(* Logix 5000 project; controller PLC_MCC1300_75F1 vendor 1 type 14 code 166 rev 32.11; software revision 32.04; part 43 of 83 *)
(* tags used below, declared in another part *)
   AUX_xDebugNewPlate : BOOL;
   CM_INPUT_Z200_Sync : CM_INPUT_Z200;
   CONST_tAux : AUX_COSTANTS;
   CONST_tPlant : UDT_PLANT_CONSTANTS;
   GP_AccTimeForGap : GP_AccTimeForGap;
   GP_TrackingAddCap : GP_TrackingAddCap;
   GP_TrackingSearchPlate : GP_TrackingSearchPlate;
   M302SpeedUp : MAC_SpeedUp;
   M302SpeedUp_ALM : MAC_SpeedUp_ALM;
   M302SpeedUp_HMR : MAC_SpeedUp_HMR;
   M302SpeedUp_tmON_ProtSnap : TIMER;
   M302SpeedUp_xFirstScanProtSnap : BOOL;
   TMP_d : DINT;
   TMP_dDebug : DINT;
   TMP_dIndex : DINT;
   TMP_dLehrSpeed : DINT;
   TMP_x : BOOL;
   xAlwaysOFF : BOOL;
   xDebugOFF : BOOL;
   Z200_SnapDataEth : UDT_ConvoyCap_ZC[2];
   Z300_BufferPlate : UDT_LINE_BUFFER_PLATE;
   Z300_Conveyor : UDT_StandConv[29];
   Z300_dEndTrackingPosition : DINT;
   Z300_LineTracking : UDT_LINE_TRACKING;
   Z301 : MAC_Zone_ML;
   Z301_HMR : MAC_Zone_ML_HMR;
(* MainProgram, continued *)

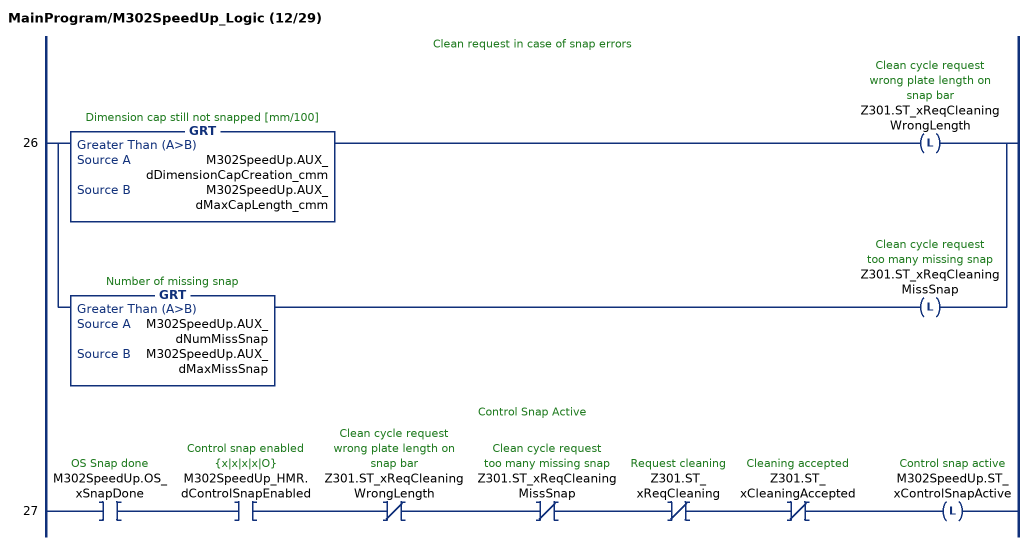
   [picture p613: MainProgram/M302SpeedUp_Logic rungs 26-27]
   // Clean request in case of snap errors
   26: [GRT(M302SpeedUp.AUX_dDimensionCapCreation_cmm,M302SpeedUp.AUX_dMaxCapLength_cmm) OTL(Z301.ST_xReqCleaningWrongLength) ,GRT(M302SpeedUp.AUX_dNumMissSnap,M302SpeedUp.AUX_dMaxMissSnap) OTL(Z301.ST_xReqCleaningMissSnap) ];
   // Control Snap Active
   27: XIC(M302SpeedUp.OS_xSnapDone)XIC(M302SpeedUp_HMR.dControlSnapEnabled)XIO(Z301.ST_xReqCleaningWrongLength)XIO(Z301.ST_xReqCleaningMissSnap)XIO(Z301.ST_xReqCleaning)XIO(Z301.ST_xCleaningAccepted)OTL(M302SpeedUp.ST_xControlSnapActive);
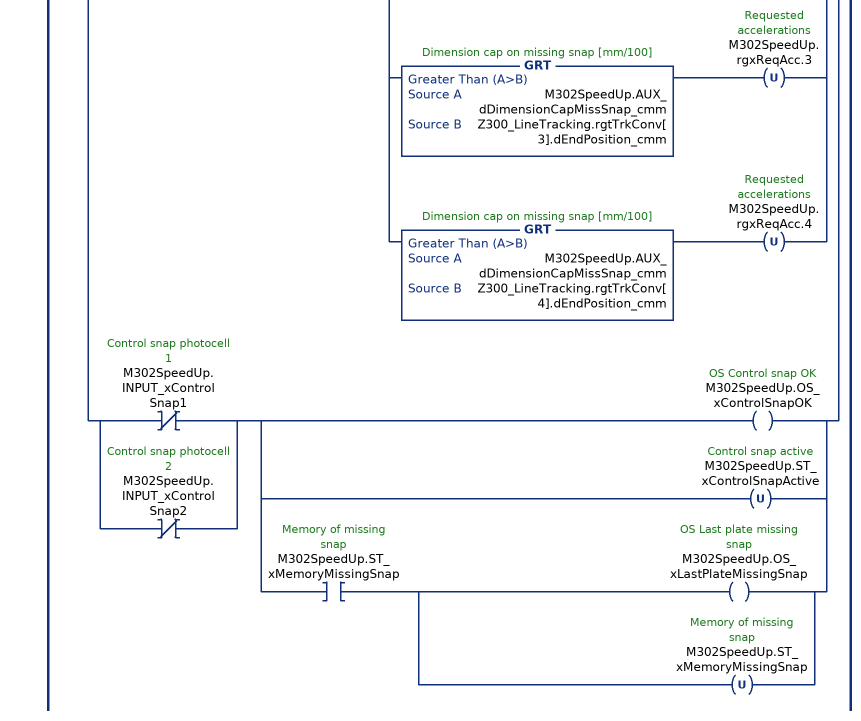
   // Missing Snap
   28: XIC(M302SpeedUp.ST_xControlSnapActive)MOV(30000,M302SpeedUp.AUX_dControlSnapLimit_cmm)[GRT(M302SpeedUp.AUX_dDimensionCapCreation_cmm,M302SpeedUp.AUX_dControlSnapLimit_cmm) [OTE(M302SpeedUp.OS_xMissingSnap) ,OTU(M302SpeedUp.ST_xControlSnapActive) ,OTU(M302SpeedUp.xReqAccAll) ,OTL(M302SpeedUp.ST_xMemoryMissingSnap) ,GRT(M302SpeedUp.AUX_dDimensionCapMissSnap_cmm,Z300_LineTracking.rgtTrkConv[0].dEndPosition_cmm) OTU(M302SpeedUp.rgxReqAcc.0) ,GRT(M302SpeedUp.AUX_dDimensionCapMissSnap_cmm,Z300_LineTracking.rgtTrkConv[1].dEndPosition_cmm) OTU(M302SpeedUp.rgxReqAcc.1) ,GRT(M302SpeedUp.AUX_dDimensionCapMissSnap_cmm,Z300_LineTracking.rgtTrkConv[2].dEndPosition_cmm) OTU(M302SpeedUp.rgxReqAcc.2) ,GRT(M302SpeedUp.AUX_dDimensionCapMissSnap_cmm,Z300_LineTracking.rgtTrkConv[3].dEndPosition_cmm) OTU(M302SpeedUp.rgxReqAcc.3) ,GRT(M302SpeedUp.AUX_dDimensionCapMissSnap_cmm,Z300_LineTracking.rgtTrkConv[4].dEndPosition_cmm) OTU(M302SpeedUp.rgxReqAcc.4) ] ,[XIO(M302SpeedUp.INPUT_xControlSnap1) ,XIO(M302SpeedUp.INPUT_xControlSnap2) ] [OTE(M302SpeedUp.OS_xControlSnapOK) ,OTU(M302SpeedUp.ST_xControlSnapActive) ,XIC(M302SpeedUp.ST_xMemoryMissingSnap) [OTE(M302SpeedUp.OS_xLastPlateMissingSnap) ,OTU(M302SpeedUp.ST_xMemoryMissingSnap) ] ] ];
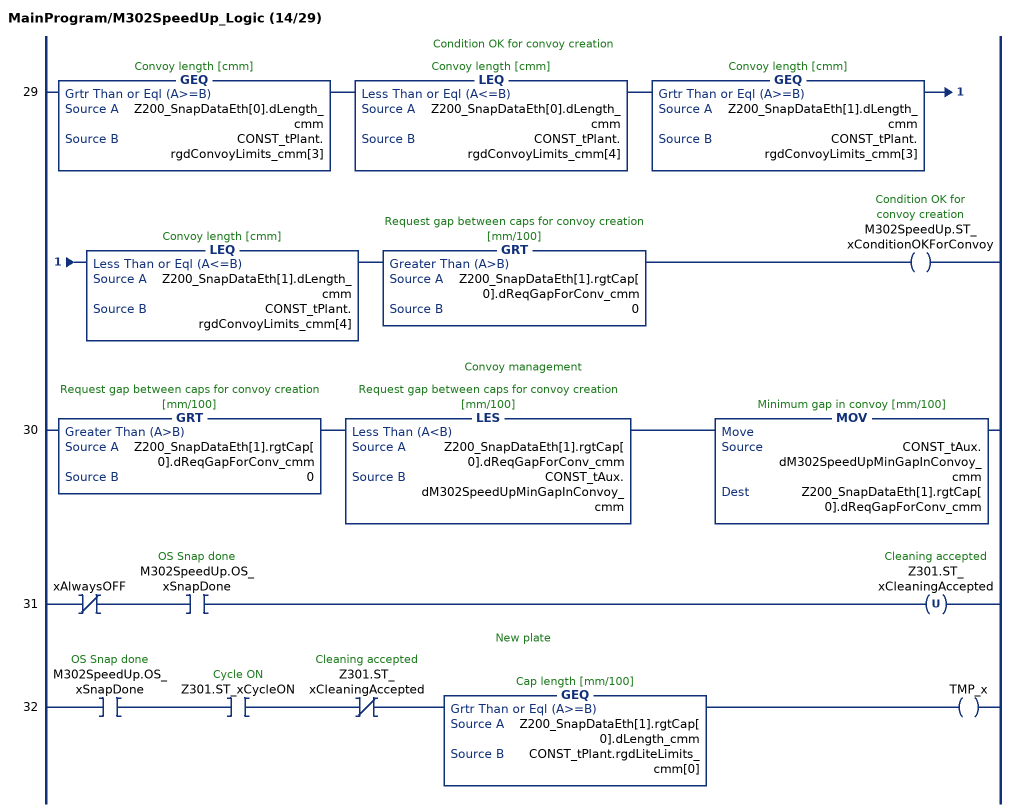
   // Condition OK for convoy creation
   29: GEQ(Z200_SnapDataEth[0].dLength_cmm,CONST_tPlant.rgdConvoyLimits_cmm[3])LEQ(Z200_SnapDataEth[0].dLength_cmm,CONST_tPlant.rgdConvoyLimits_cmm[4])GEQ(Z200_SnapDataEth[1].dLength_cmm,CONST_tPlant.rgdConvoyLimits_cmm[3])LEQ(Z200_SnapDataEth[1].dLength_cmm,CONST_tPlant.rgdConvoyLimits_cmm[4])GRT(Z200_SnapDataEth[1].rgtCap[0].dReqGapForConv_cmm,0)OTE(M302SpeedUp.ST_xConditionOKForConvoy);
   // Convoy management
   30: GRT(Z200_SnapDataEth[1].rgtCap[0].dReqGapForConv_cmm,0)LES(Z200_SnapDataEth[1].rgtCap[0].dReqGapForConv_cmm,CONST_tAux.dM302SpeedUpMinGapInConvoy_cmm)MOV(CONST_tAux.dM302SpeedUpMinGapInConvoy_cmm,Z200_SnapDataEth[1].rgtCap[0].dReqGapForConv_cmm);
   31: XIO(xAlwaysOFF)XIC(M302SpeedUp.OS_xSnapDone)OTU(Z301.ST_xCleaningAccepted);
   // New plate
   32: XIC(M302SpeedUp.OS_xSnapDone)XIC(Z301.ST_xCycleON)XIO(Z301.ST_xCleaningAccepted)GEQ(Z200_SnapDataEth[1].rgtCap[0].dLength_cmm,CONST_tPlant.rgdLiteLimits_cmm[0])OTE(TMP_x);
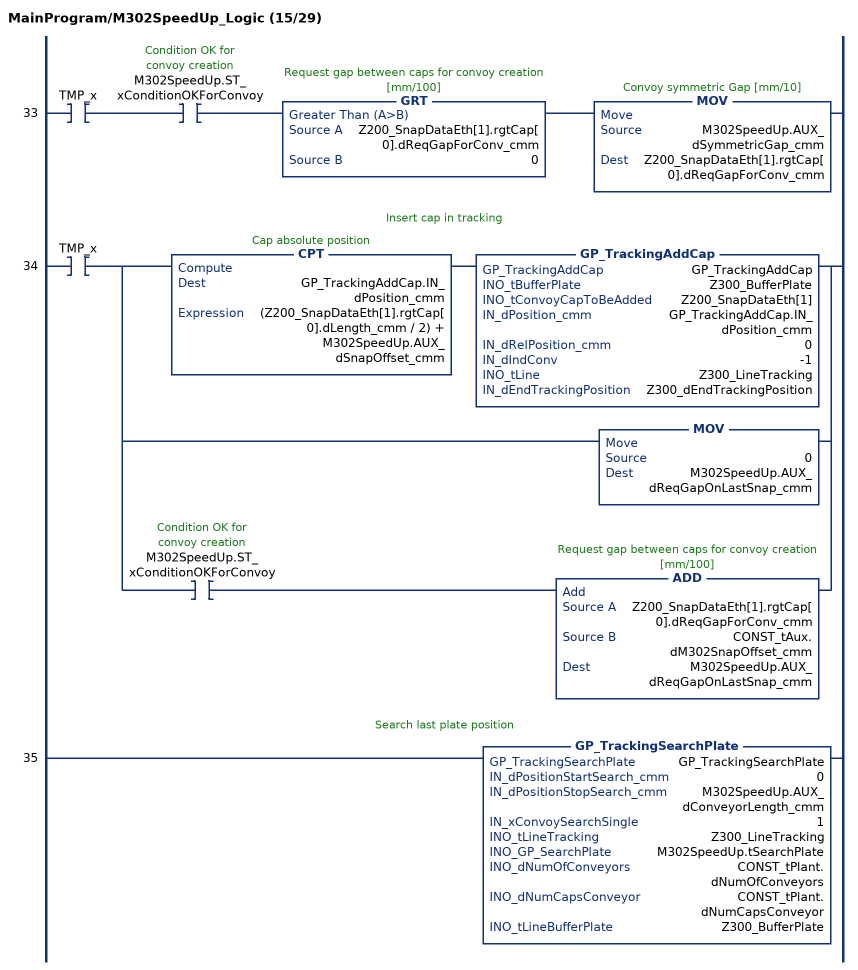
   33: XIC(TMP_x)XIC(M302SpeedUp.ST_xConditionOKForConvoy)GRT(Z200_SnapDataEth[1].rgtCap[0].dReqGapForConv_cmm,0)MOV(M302SpeedUp.AUX_dSymmetricGap_cmm,Z200_SnapDataEth[1].rgtCap[0].dReqGapForConv_cmm);
   // Insert cap in tracking
   34: XIC(TMP_x)[CPT(GP_TrackingAddCap.IN_dPosition_cmm,(Z200_SnapDataEth[1].rgtCap[0].dLength_cmm / 2) + M302SpeedUp.AUX_dSnapOffset_cmm) GP_TrackingAddCap(GP_TrackingAddCap,Z300_BufferPlate,Z200_SnapDataEth[1],GP_TrackingAddCap.IN_dPosition_cmm,0,-1,Z300_LineTracking,Z300_dEndTrackingPosition) ,MOV(0,M302SpeedUp.AUX_dReqGapOnLastSnap_cmm) ,XIC(M302SpeedUp.ST_xConditionOKForConvoy) ADD(Z200_SnapDataEth[1].rgtCap[0].dReqGapForConv_cmm,CONST_tAux.dM302SnapOffset_cmm,M302SpeedUp.AUX_dReqGapOnLastSnap_cmm) ];
   // Search last plate position
   35: GP_TrackingSearchPlate(GP_TrackingSearchPlate,0,M302SpeedUp.AUX_dConveyorLength_cmm,1,Z300_LineTracking,M302SpeedUp.tSearchPlate,CONST_tPlant.dNumOfConveyors,CONST_tPlant.dNumCapsConveyor,Z300_BufferPlate);
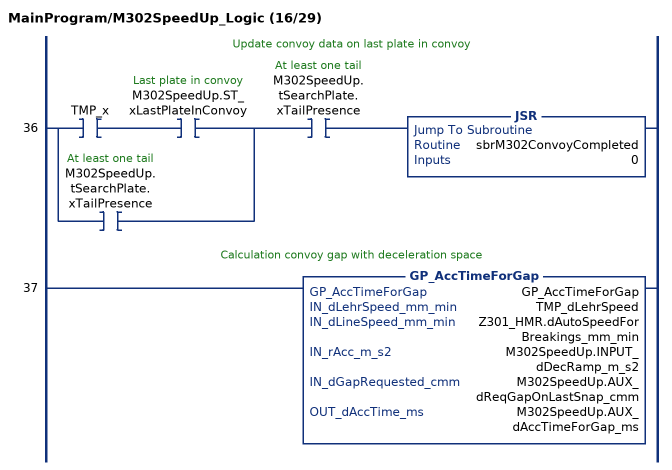
   // Update convoy data on last plate in convoy
   36: [XIC(TMP_x) XIC(M302SpeedUp.ST_xLastPlateInConvoy) ,XIC(M302SpeedUp.tSearchPlate.xTailPresence) ]XIC(M302SpeedUp.tSearchPlate.xTailPresence)JSR(sbrM302ConvoyCompleted,0);
   // Calculation convoy gap with deceleration space
   37: GP_AccTimeForGap(GP_AccTimeForGap,TMP_dLehrSpeed,Z301_HMR.dAutoSpeedForBreakings_mm_min,M302SpeedUp.INPUT_dDecRamp_m_s2,M302SpeedUp.AUX_dReqGapOnLastSnap_cmm,M302SpeedUp.AUX_dAccTimeForGap_ms);
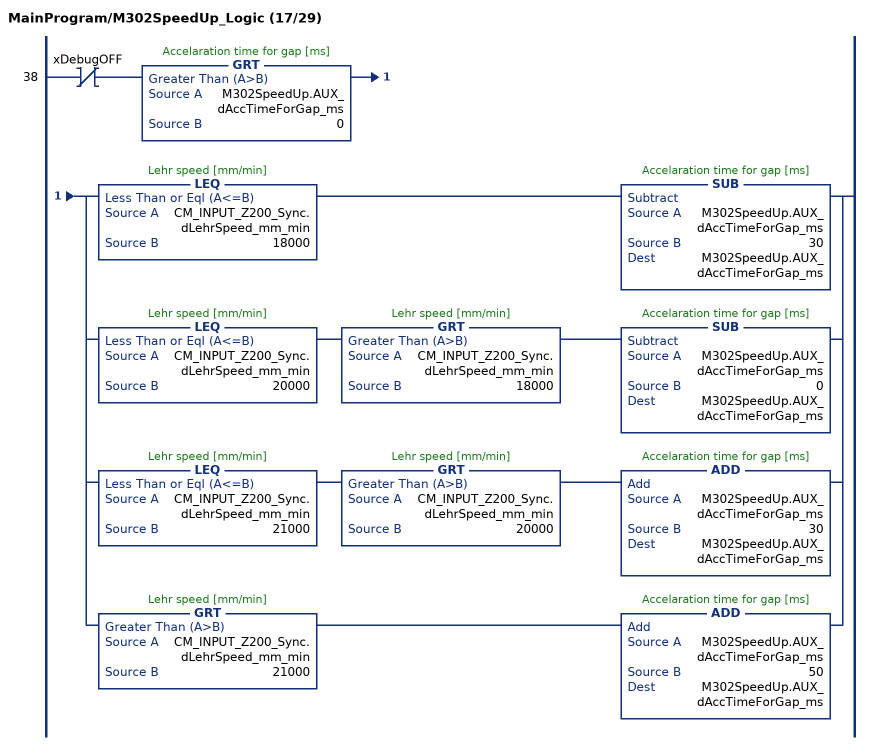
   38: XIO(xDebugOFF)GRT(M302SpeedUp.AUX_dAccTimeForGap_ms,0)[LEQ(CM_INPUT_Z200_Sync.dLehrSpeed_mm_min,18000) SUB(M302SpeedUp.AUX_dAccTimeForGap_ms,30,M302SpeedUp.AUX_dAccTimeForGap_ms) ,LEQ(CM_INPUT_Z200_Sync.dLehrSpeed_mm_min,20000) GRT(CM_INPUT_Z200_Sync.dLehrSpeed_mm_min,18000) SUB(M302SpeedUp.AUX_dAccTimeForGap_ms,0,M302SpeedUp.AUX_dAccTimeForGap_ms) ,LEQ(CM_INPUT_Z200_Sync.dLehrSpeed_mm_min,21000) GRT(CM_INPUT_Z200_Sync.dLehrSpeed_mm_min,20000) ADD(M302SpeedUp.AUX_dAccTimeForGap_ms,30,M302SpeedUp.AUX_dAccTimeForGap_ms) ,GRT(CM_INPUT_Z200_Sync.dLehrSpeed_mm_min,21000) ADD(M302SpeedUp.AUX_dAccTimeForGap_ms,50,M302SpeedUp.AUX_dAccTimeForGap_ms) ];
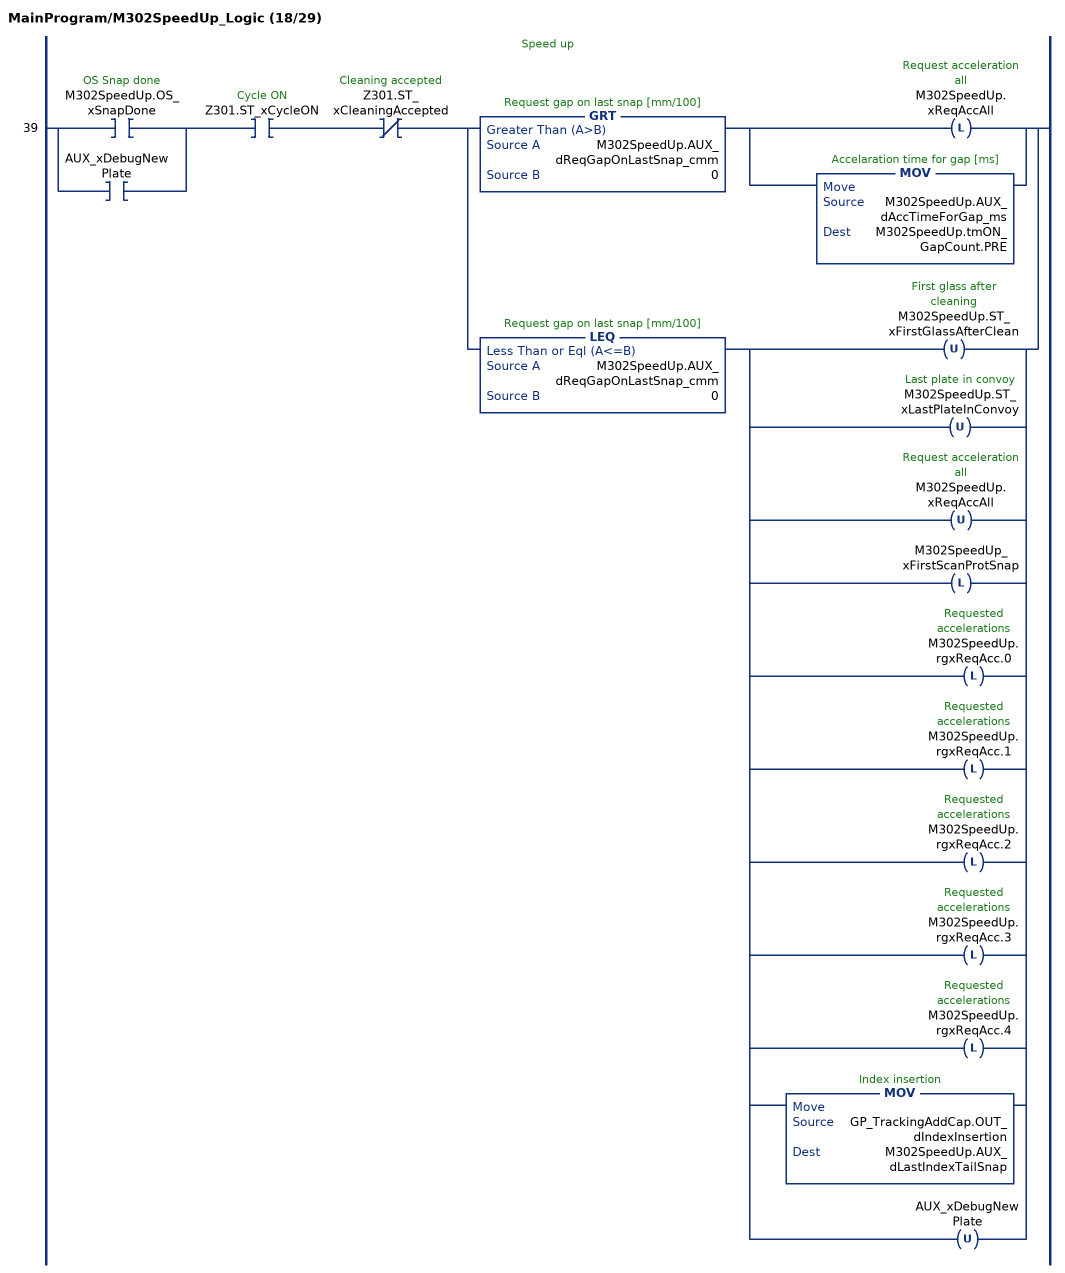
   // Speed up
   39: [XIC(M302SpeedUp.OS_xSnapDone) ,XIC(AUX_xDebugNewPlate) ]XIC(Z301.ST_xCycleON)XIO(Z301.ST_xCleaningAccepted)[GRT(M302SpeedUp.AUX_dReqGapOnLastSnap_cmm,0) [OTL(M302SpeedUp.xReqAccAll) ,MOV(M302SpeedUp.AUX_dAccTimeForGap_ms,M302SpeedUp.tmON_GapCount.PRE) ] ,LEQ(M302SpeedUp.AUX_dReqGapOnLastSnap_cmm,0) [OTU(M302SpeedUp.ST_xFirstGlassAfterClean) ,OTU(M302SpeedUp.ST_xLastPlateInConvoy) ,OTU(M302SpeedUp.xReqAccAll) ,OTL(M302SpeedUp_xFirstScanProtSnap) ,OTL(M302SpeedUp.rgxReqAcc.0) ,OTL(M302SpeedUp.rgxReqAcc.1) ,OTL(M302SpeedUp.rgxReqAcc.2) ,OTL(M302SpeedUp.rgxReqAcc.3) ,OTL(M302SpeedUp.rgxReqAcc.4) ,MOV(GP_TrackingAddCap.OUT_dIndexInsertion,M302SpeedUp.AUX_dLastIndexTailSnap) ,OTU(AUX_xDebugNewPlate) ] ];
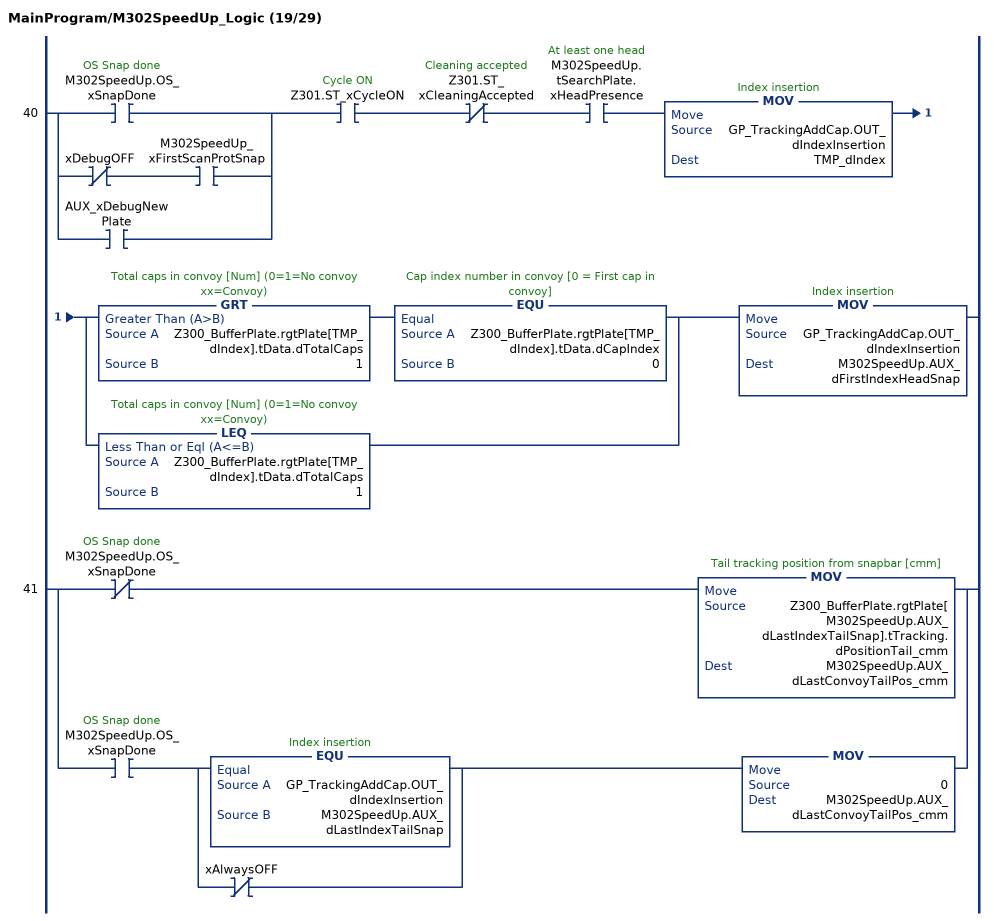
   40: [XIC(M302SpeedUp.OS_xSnapDone) ,XIO(xDebugOFF) XIC(M302SpeedUp_xFirstScanProtSnap) ,XIC(AUX_xDebugNewPlate) ]XIC(Z301.ST_xCycleON)XIO(Z301.ST_xCleaningAccepted)XIC(M302SpeedUp.tSearchPlate.xHeadPresence)MOV(GP_TrackingAddCap.OUT_dIndexInsertion,TMP_dIndex)[GRT(Z300_BufferPlate.rgtPlate[TMP_dIndex].tData.dTotalCaps,1) EQU(Z300_BufferPlate.rgtPlate[TMP_dIndex].tData.dCapIndex,0) ,LEQ(Z300_BufferPlate.rgtPlate[TMP_dIndex].tData.dTotalCaps,1) ]MOV(GP_TrackingAddCap.OUT_dIndexInsertion,M302SpeedUp.AUX_dFirstIndexHeadSnap);
   41: [XIO(M302SpeedUp.OS_xSnapDone) MOV(Z300_BufferPlate.rgtPlate[M302SpeedUp.AUX_dLastIndexTailSnap].tTracking.dPositionTail_cmm,M302SpeedUp.AUX_dLastConvoyTailPos_cmm) ,XIC(M302SpeedUp.OS_xSnapDone) [EQU(GP_TrackingAddCap.OUT_dIndexInsertion,M302SpeedUp.AUX_dLastIndexTailSnap) ,XIO(xAlwaysOFF) ] MOV(0,M302SpeedUp.AUX_dLastConvoyTailPos_cmm) ];
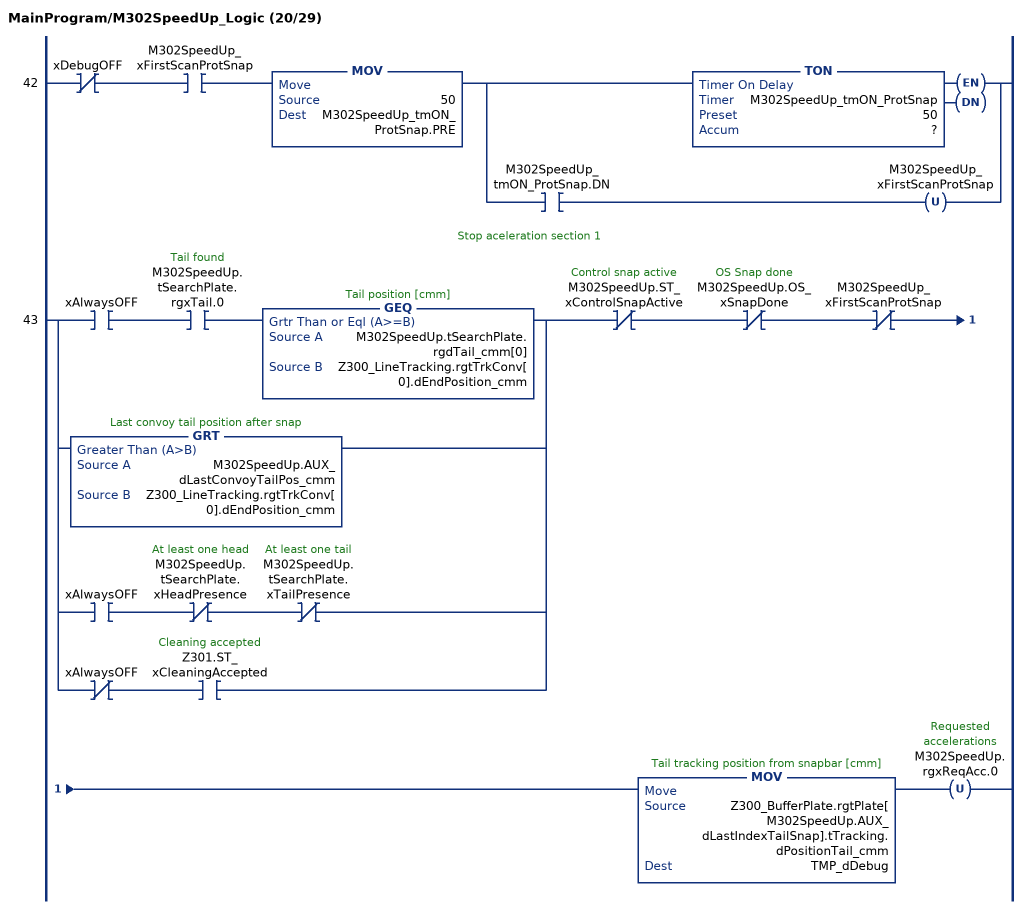
   42: XIO(xDebugOFF)XIC(M302SpeedUp_xFirstScanProtSnap)MOV(50,M302SpeedUp_tmON_ProtSnap.PRE)[TON(M302SpeedUp_tmON_ProtSnap,?,?) ,XIC(M302SpeedUp_tmON_ProtSnap.DN) OTU(M302SpeedUp_xFirstScanProtSnap) ];
   // Stop aceleration section 1
   43: [[XIC(xAlwaysOFF) XIC(M302SpeedUp.tSearchPlate.rgxTail.0) GEQ(M302SpeedUp.tSearchPlate.rgdTail_cmm[0],Z300_LineTracking.rgtTrkConv[0].dEndPosition_cmm) ,GRT(M302SpeedUp.AUX_dLastConvoyTailPos_cmm,Z300_LineTracking.rgtTrkConv[0].dEndPosition_cmm) ] ,XIC(xAlwaysOFF) XIO(M302SpeedUp.tSearchPlate.xHeadPresence) XIO(M302SpeedUp.tSearchPlate.xTailPresence) ,XIO(xAlwaysOFF) XIC(Z301.ST_xCleaningAccepted) ]XIO(M302SpeedUp.ST_xControlSnapActive)XIO(M302SpeedUp.OS_xSnapDone)XIO(M302SpeedUp_xFirstScanProtSnap)MOV(Z300_BufferPlate.rgtPlate[M302SpeedUp.AUX_dLastIndexTailSnap].tTracking.dPositionTail_cmm,TMP_dDebug)OTU(M302SpeedUp.rgxReqAcc.0);
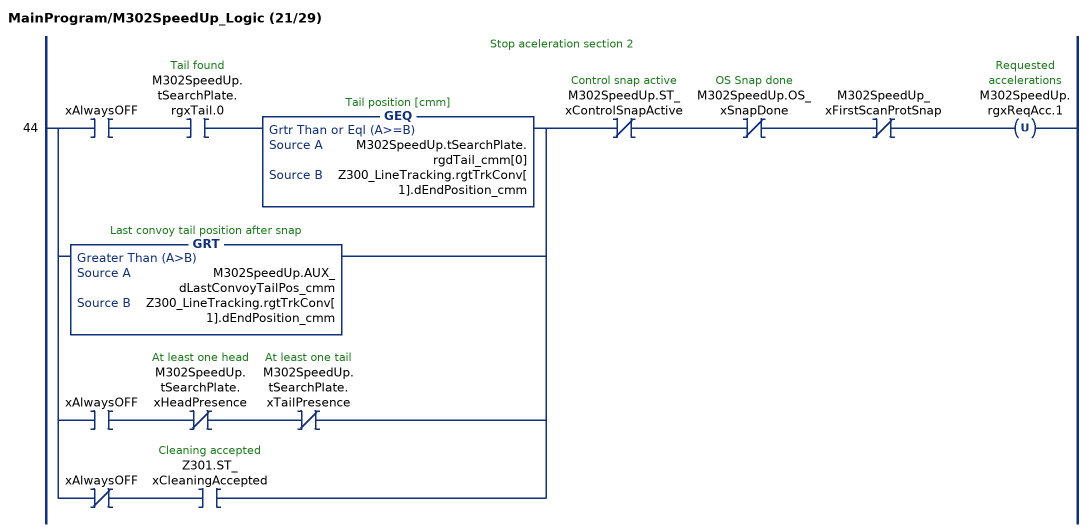
   // Stop aceleration section 2
   44: [[XIC(xAlwaysOFF) XIC(M302SpeedUp.tSearchPlate.rgxTail.0) GEQ(M302SpeedUp.tSearchPlate.rgdTail_cmm[0],Z300_LineTracking.rgtTrkConv[1].dEndPosition_cmm) ,GRT(M302SpeedUp.AUX_dLastConvoyTailPos_cmm,Z300_LineTracking.rgtTrkConv[1].dEndPosition_cmm) ] ,XIC(xAlwaysOFF) XIO(M302SpeedUp.tSearchPlate.xHeadPresence) XIO(M302SpeedUp.tSearchPlate.xTailPresence) ,XIO(xAlwaysOFF) XIC(Z301.ST_xCleaningAccepted) ]XIO(M302SpeedUp.ST_xControlSnapActive)XIO(M302SpeedUp.OS_xSnapDone)XIO(M302SpeedUp_xFirstScanProtSnap)OTU(M302SpeedUp.rgxReqAcc.1);
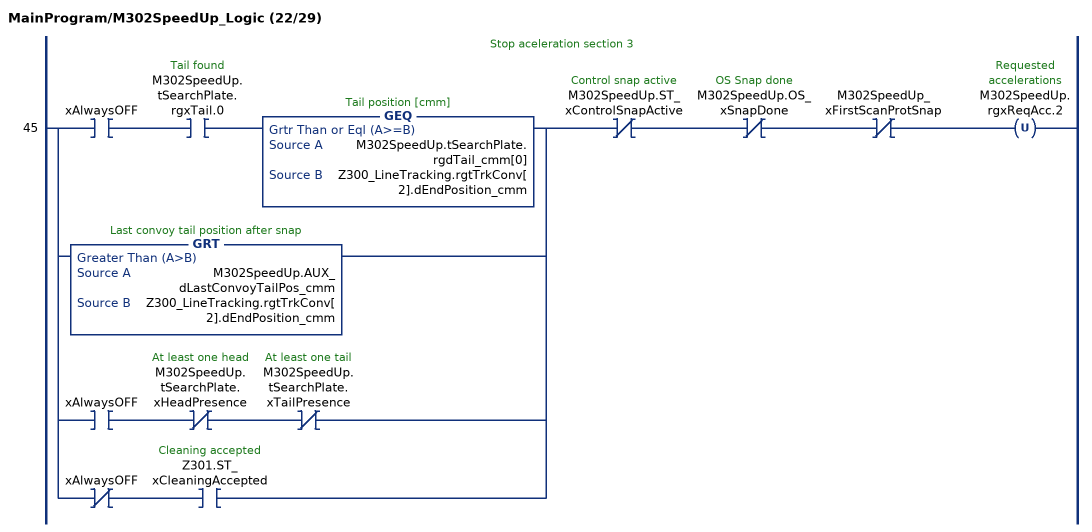
   // Stop aceleration section 3
   45: [[XIC(xAlwaysOFF) XIC(M302SpeedUp.tSearchPlate.rgxTail.0) GEQ(M302SpeedUp.tSearchPlate.rgdTail_cmm[0],Z300_LineTracking.rgtTrkConv[2].dEndPosition_cmm) ,GRT(M302SpeedUp.AUX_dLastConvoyTailPos_cmm,Z300_LineTracking.rgtTrkConv[2].dEndPosition_cmm) ] ,XIC(xAlwaysOFF) XIO(M302SpeedUp.tSearchPlate.xHeadPresence) XIO(M302SpeedUp.tSearchPlate.xTailPresence) ,XIO(xAlwaysOFF) XIC(Z301.ST_xCleaningAccepted) ]XIO(M302SpeedUp.ST_xControlSnapActive)XIO(M302SpeedUp.OS_xSnapDone)XIO(M302SpeedUp_xFirstScanProtSnap)OTU(M302SpeedUp.rgxReqAcc.2);
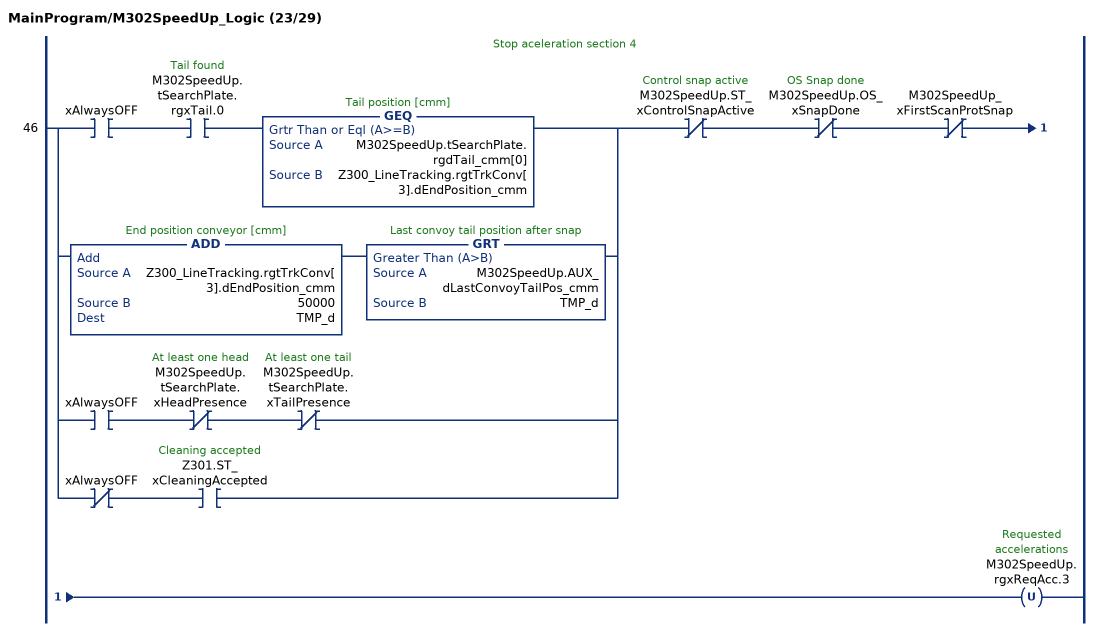
   // Stop aceleration section 4
   46: [[XIC(xAlwaysOFF) XIC(M302SpeedUp.tSearchPlate.rgxTail.0) GEQ(M302SpeedUp.tSearchPlate.rgdTail_cmm[0],Z300_LineTracking.rgtTrkConv[3].dEndPosition_cmm) ,ADD(Z300_LineTracking.rgtTrkConv[3].dEndPosition_cmm,50000,TMP_d) GRT(M302SpeedUp.AUX_dLastConvoyTailPos_cmm,TMP_d) ] ,XIC(xAlwaysOFF) XIO(M302SpeedUp.tSearchPlate.xHeadPresence) XIO(M302SpeedUp.tSearchPlate.xTailPresence) ,XIO(xAlwaysOFF) XIC(Z301.ST_xCleaningAccepted) ]XIO(M302SpeedUp.ST_xControlSnapActive)XIO(M302SpeedUp.OS_xSnapDone)XIO(M302SpeedUp_xFirstScanProtSnap)OTU(M302SpeedUp.rgxReqAcc.3);
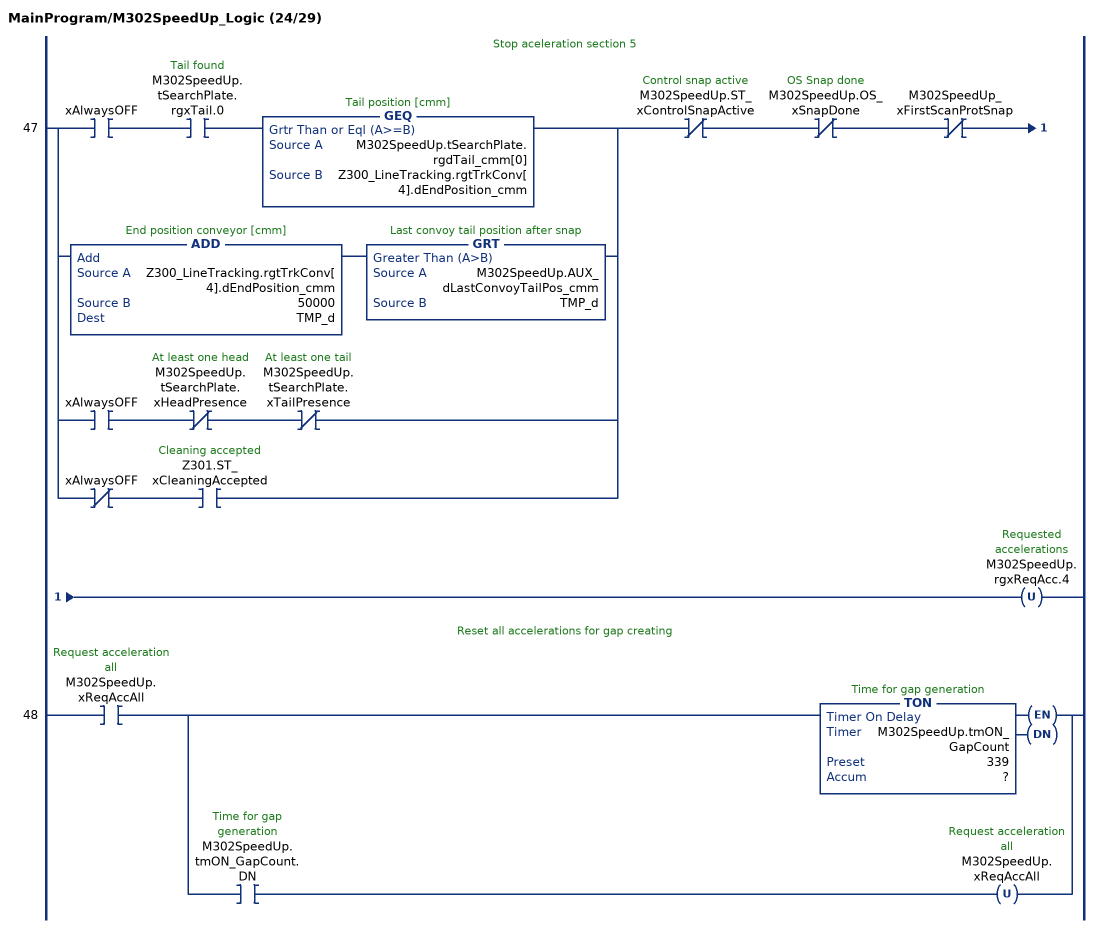
   // Stop aceleration section 5
   47: [[XIC(xAlwaysOFF) XIC(M302SpeedUp.tSearchPlate.rgxTail.0) GEQ(M302SpeedUp.tSearchPlate.rgdTail_cmm[0],Z300_LineTracking.rgtTrkConv[4].dEndPosition_cmm) ,ADD(Z300_LineTracking.rgtTrkConv[4].dEndPosition_cmm,50000,TMP_d) GRT(M302SpeedUp.AUX_dLastConvoyTailPos_cmm,TMP_d) ] ,XIC(xAlwaysOFF) XIO(M302SpeedUp.tSearchPlate.xHeadPresence) XIO(M302SpeedUp.tSearchPlate.xTailPresence) ,XIO(xAlwaysOFF) XIC(Z301.ST_xCleaningAccepted) ]XIO(M302SpeedUp.ST_xControlSnapActive)XIO(M302SpeedUp.OS_xSnapDone)XIO(M302SpeedUp_xFirstScanProtSnap)OTU(M302SpeedUp.rgxReqAcc.4);
   // Reset all accelerations for gap creating
   48: XIC(M302SpeedUp.xReqAccAll)[TON(M302SpeedUp.tmON_GapCount,?,?) ,XIC(M302SpeedUp.tmON_GapCount.DN) OTU(M302SpeedUp.xReqAccAll) ];
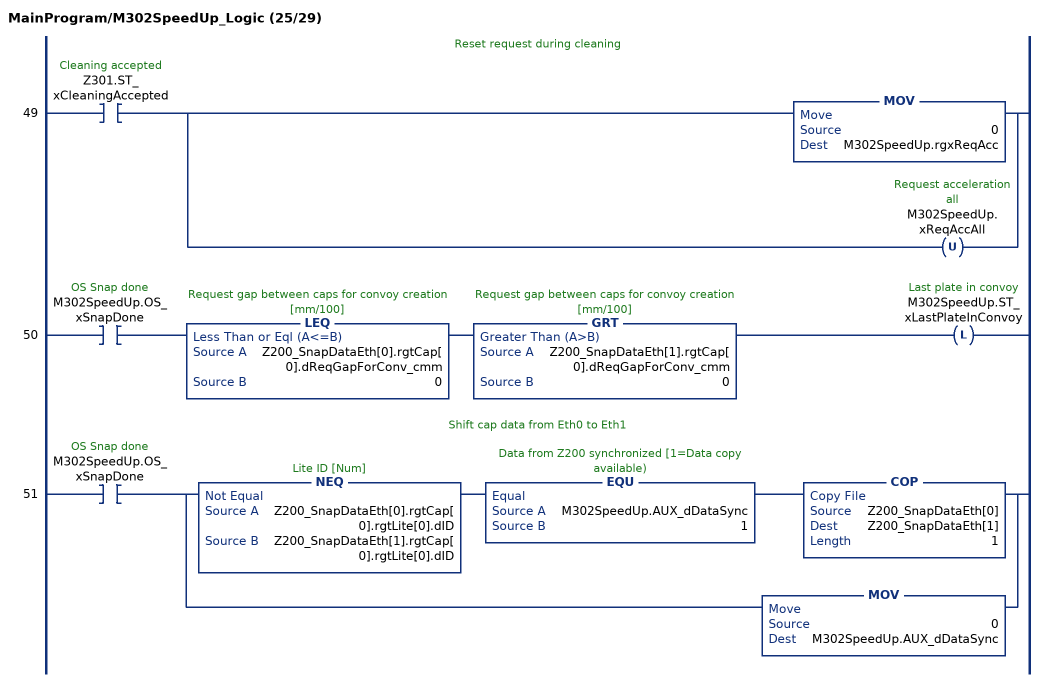
   // Reset request during cleaning
   49: XIC(Z301.ST_xCleaningAccepted)[MOV(0,M302SpeedUp.rgxReqAcc) ,OTU(M302SpeedUp.xReqAccAll) ];
   50: XIC(M302SpeedUp.OS_xSnapDone)LEQ(Z200_SnapDataEth[0].rgtCap[0].dReqGapForConv_cmm,0)GRT(Z200_SnapDataEth[1].rgtCap[0].dReqGapForConv_cmm,0)OTL(M302SpeedUp.ST_xLastPlateInConvoy);
   // Shift cap data from Eth0 to Eth1
   51: XIC(M302SpeedUp.OS_xSnapDone)[NEQ(Z200_SnapDataEth[0].rgtCap[0].rgtLite[0].dID,Z200_SnapDataEth[1].rgtCap[0].rgtLite[0].dID) EQU(M302SpeedUp.AUX_dDataSync,1) COP(Z200_SnapDataEth[0],Z200_SnapDataEth[1],1) ,MOV(0,M302SpeedUp.AUX_dDataSync) ];
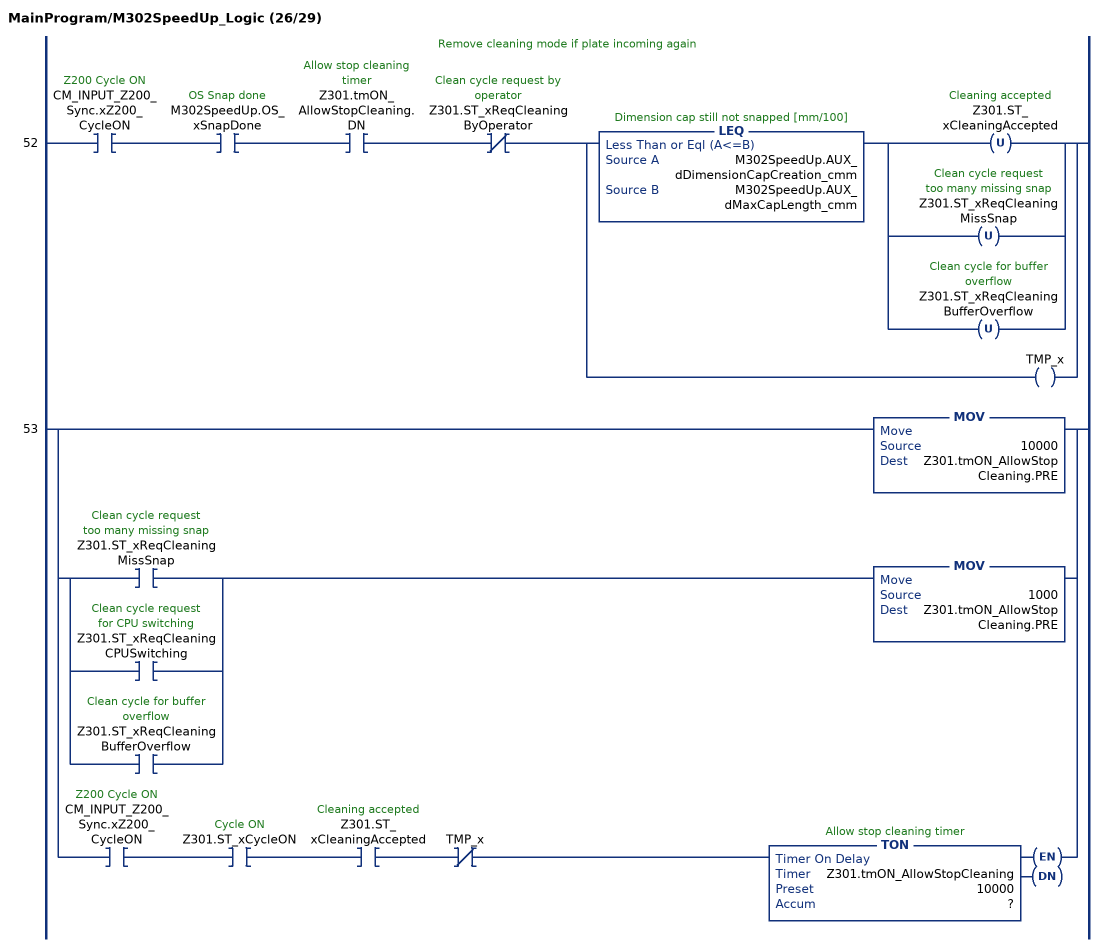
   // Remove cleaning mode if plate incoming again
   52: XIC(CM_INPUT_Z200_Sync.xZ200_CycleON)XIC(M302SpeedUp.OS_xSnapDone)XIC(Z301.tmON_AllowStopCleaning.DN)XIO(Z301.ST_xReqCleaningByOperator)[LEQ(M302SpeedUp.AUX_dDimensionCapCreation_cmm,M302SpeedUp.AUX_dMaxCapLength_cmm) [OTU(Z301.ST_xCleaningAccepted) ,[OTU(Z301.ST_xReqCleaningMissSnap) ,OTU(Z301.ST_xReqCleaningBufferOverflow) ] ] ,OTE(TMP_x) ];
   53: [MOV(10000,Z301.tmON_AllowStopCleaning.PRE) ,[XIC(Z301.ST_xReqCleaningMissSnap) ,XIC(Z301.ST_xReqCleaningCPUSwitching) ,XIC(Z301.ST_xReqCleaningBufferOverflow) ] MOV(1000,Z301.tmON_AllowStopCleaning.PRE) ,XIC(CM_INPUT_Z200_Sync.xZ200_CycleON) XIC(Z301.ST_xCycleON) XIC(Z301.ST_xCleaningAccepted) XIO(TMP_x) TON(Z301.tmON_AllowStopCleaning,?,?) ];
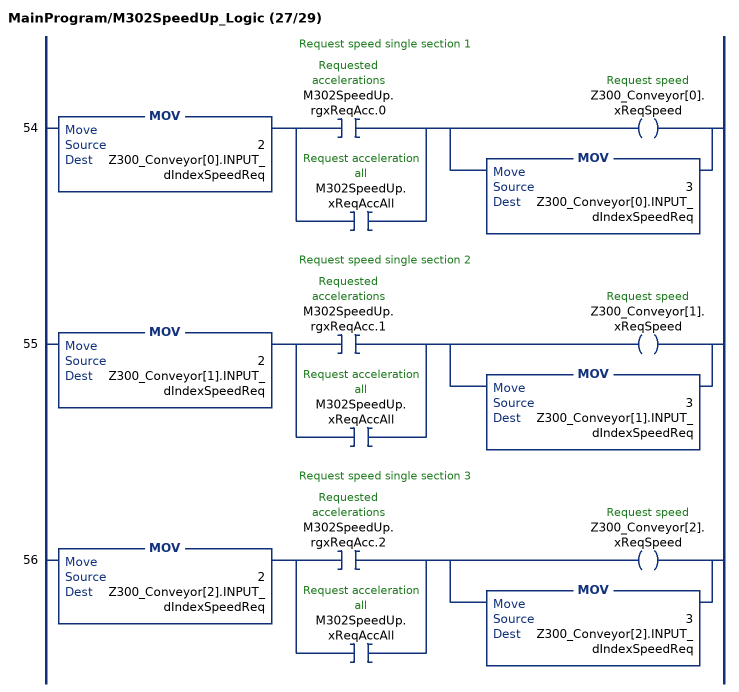
   // Request speed single section 1
   54: MOV(2,Z300_Conveyor[0].INPUT_dIndexSpeedReq)[XIC(M302SpeedUp.rgxReqAcc.0) ,XIC(M302SpeedUp.xReqAccAll) ][OTE(Z300_Conveyor[0].xReqSpeed) ,MOV(3,Z300_Conveyor[0].INPUT_dIndexSpeedReq) ];
   // Request speed single section 2
   55: MOV(2,Z300_Conveyor[1].INPUT_dIndexSpeedReq)[XIC(M302SpeedUp.rgxReqAcc.1) ,XIC(M302SpeedUp.xReqAccAll) ][OTE(Z300_Conveyor[1].xReqSpeed) ,MOV(3,Z300_Conveyor[1].INPUT_dIndexSpeedReq) ];
   // Request speed single section 3
   56: MOV(2,Z300_Conveyor[2].INPUT_dIndexSpeedReq)[XIC(M302SpeedUp.rgxReqAcc.2) ,XIC(M302SpeedUp.xReqAccAll) ][OTE(Z300_Conveyor[2].xReqSpeed) ,MOV(3,Z300_Conveyor[2].INPUT_dIndexSpeedReq) ];
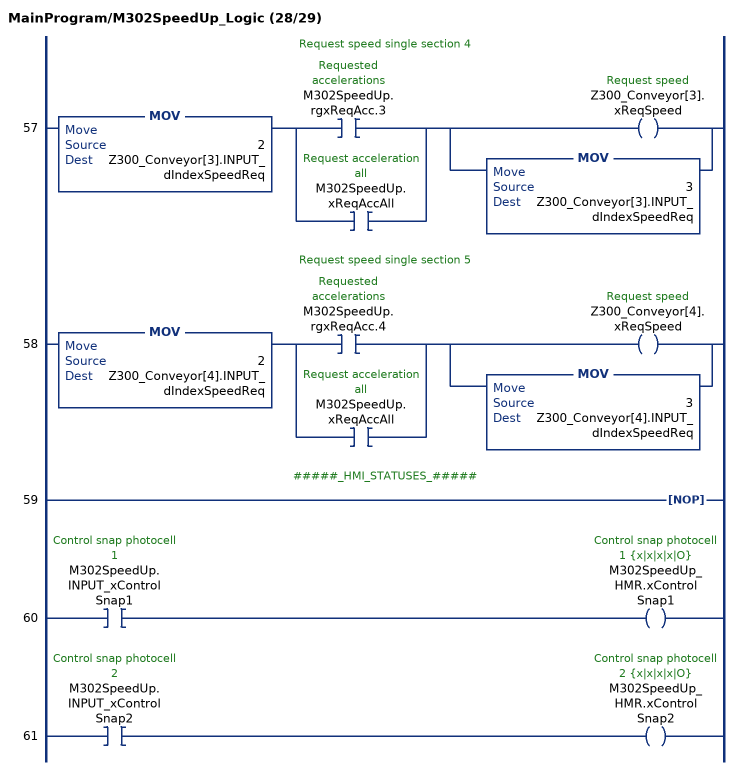
   // Request speed single section 4
   57: MOV(2,Z300_Conveyor[3].INPUT_dIndexSpeedReq)[XIC(M302SpeedUp.rgxReqAcc.3) ,XIC(M302SpeedUp.xReqAccAll) ][OTE(Z300_Conveyor[3].xReqSpeed) ,MOV(3,Z300_Conveyor[3].INPUT_dIndexSpeedReq) ];
   // Request speed single section 5
   58: MOV(2,Z300_Conveyor[4].INPUT_dIndexSpeedReq)[XIC(M302SpeedUp.rgxReqAcc.4) ,XIC(M302SpeedUp.xReqAccAll) ][OTE(Z300_Conveyor[4].xReqSpeed) ,MOV(3,Z300_Conveyor[4].INPUT_dIndexSpeedReq) ];
   // #####_HMI_STATUSES_#####
   59: NOP();
   60: XIC(M302SpeedUp.INPUT_xControlSnap1)OTE(M302SpeedUp_HMR.xControlSnap1);
   61: XIC(M302SpeedUp.INPUT_xControlSnap2)OTE(M302SpeedUp_HMR.xControlSnap2);
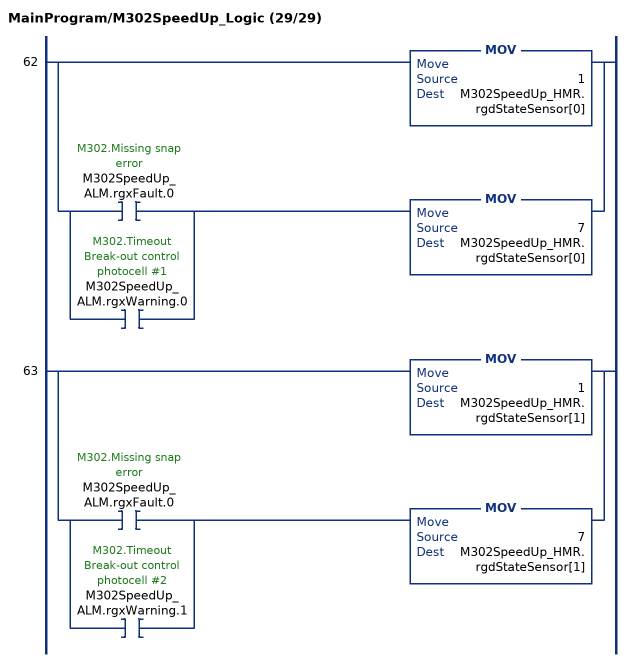
   62: [MOV(1,M302SpeedUp_HMR.rgdStateSensor[0]) ,[XIC(M302SpeedUp_ALM.rgxFault.0) ,XIC(M302SpeedUp_ALM.rgxWarning.0) ] MOV(7,M302SpeedUp_HMR.rgdStateSensor[0]) ];
   63: [MOV(1,M302SpeedUp_HMR.rgdStateSensor[1]) ,[XIC(M302SpeedUp_ALM.rgxFault.0) ,XIC(M302SpeedUp_ALM.rgxWarning.1) ] MOV(7,M302SpeedUp_HMR.rgdStateSensor[1]) ];
END_ROUTINE
